   "Carrier_67_SitopSelectStatus" AT %I3716.3 : Bool;   // SITOP SELECT STATUS
   "Carrier_67_DCsupplyOnPSCB2" AT %I3716.4 : Bool;   // DC SUPPLY ON PSCB 2
   "Carrier_67_SpareInput(4_5)" AT %I3716.5 : Bool;   // SPARE INPUT
   "Carrier_67_SpareInput(4_6)" AT %I3716.6 : Bool;   // SPARE INPUT
   "Carrier_67_SpareInput(4_7)" AT %I3716.7 : Bool;   // SPARE INPUT
   "Carrier_67_PB1_ProdHoldLH" AT %I3717.0 : Bool;   // PB 1 PRODUCTION HOLD LH
   "Carrier_67_PB2_ResetLH" AT %I3717.1 : Bool;   // PB 2 RESET LH
   "Carrier_67_PB3_ProdHoldRH" AT %I3717.2 : Bool;   // PB 3 PRODUCTION HOLD RH
   "Carrier_67_PB4_ResetRH" AT %I3717.3 : Bool;   // PB 4 RESET RH
   "Carrier_67_SpareInput(4_14)" AT %I3717.4 : Bool;   // SPARE INPUT
   "Carrier_67_SpareInput(4_15)" AT %I3717.5 : Bool;   // SPARE INPUT
   "Carrier_67_SpareInput(4_16)" AT %I3717.6 : Bool;   // SPARE INPUT
   "Carrier_67_SpareInput(4_17)" AT %I3717.7 : Bool;   // SPARE INPUT
   "Carrier_67_Slot5_Output" AT %IW3718 : Word;   // SLOT 5 OUTPUT WORD
   "Carrier_67_IRD400_HMI_24VDC_ENABLE" AT %I3718.0 : Bool;   // IRD 400 PANEL HMI 24V DC POWER
   "Carrier_67_FaultLight_LH" AT %I3718.1 : Bool;   // FAULT LIGHT LH
   "Carrier_67_RunLight_LH" AT %I3718.2 : Bool;   // RUN LIGHT LH
   "Carrier_67_FaultLight_RH" AT %I3718.3 : Bool;   // FAULT LIGHT RH
   "Carrier_67_RunLight_RH" AT %I3718.4 : Bool;   // RUN LIGHT RH
   "Carrier_67_SpareOutput(5_5)" AT %I3718.5 : Bool;   // SPARE OUTPUT
   "Carrier_67_SpareOutput(5_6)" AT %I3718.6 : Bool;   // SPARE OUTPUT
   "Carrier_67_SpareOutput(5_7)" AT %I3718.7 : Bool;   // SPARE OUTPUT
   "Carrier_67_ActualSpeed" AT %IW3720 : Word;   // ACTUAL SPEED
   "Carrier_67_CarrierDriveAlarm" AT %IW3722 : Word;   // CARRIER DRIVE ALARM
   "Carrier_67_CarrierDriveWarning" AT %IW3724 : Word;   // CARRIER DRIVE WARNING
   "Carrier_68_Status" AT %IW3750 : Word;   // CARRIER STATUS WORD
   "Carrier_68_Status.0" AT %I3750.0 : Bool;   // HEARTBEAT
   "Carrier_68_Status.1" AT %I3750.1 : Bool;   // MANUAL
   "Carrier_68_Status.2" AT %I3750.2 : Bool;   // IN_AUTO
   "Carrier_68_Status.3" AT %I3750.3 : Bool;   // POSITIONING_COMPLETE
   "Carrier_68_Status.4" AT %I3750.4 : Bool;   // PRODUCTION HOLD
   "Carrier_68_Status.5" AT %I3750.5 : Bool;   // CARRIER MOVING FORWARD
   "Carrier_68_Status.6" AT %I3750.6 : Bool;   // CARRIER MOVING REVERSE
   "Carrier_68_Status.7" AT %I3750.7 : Bool;   // CARRIER FAULT
   "Carrier_68_Status.8" AT %I3751.0 : Bool;   // CRASH DETECT TRIPPED
   "Carrier_68_Status.9" AT %I3751.1 : Bool;
   "Carrier_68_Status.10" AT %I3751.2 : Bool;
   "Carrier_68_Status.11" AT %I3751.3 : Bool;
   "Carrier_68_Status.12" AT %I3751.4 : Bool;
   "Carrier_68_Status.13" AT %I3751.5 : Bool;
   "Carrier_68_Status.14" AT %I3751.6 : Bool;
   "Carrier_68_Status.15" AT %I3751.7 : Bool;
   "Carrier_68_SDCFaultCode" AT %IW3752 : Word;   // SDC FAULT CODE
   "Carrier_68_CarrierPosition" AT %ID3754 : DWord;   // CARRIER POSITION
   "Carrier_68_CarrierNumber" AT %IW3758 : Word;   // CARRIER NUMBER
   "Carrier_68_G120DControlWord" AT %IW3760 : Word;   // G120D_STW1_CONTROL
   "Carrier_68_G120DControlWord.0" AT %I3760.0 : Bool;   // Bit_00_ON
   "Carrier_68_G120DControlWord.1" AT %I3760.1 : Bool;   // Bit_01_AUS2_INH
   "Carrier_68_G120DControlWord.2" AT %I3760.2 : Bool;   // Bit_02_AUS3_STOP
   "Carrier_68_G120DControlWord.3" AT %I3760.3 : Bool;   // Bit_03_EN
   "Carrier_68_G120DControlWord.4" AT %I3760.4 : Bool;   // Bit_04_EN_RAMP
   "Carrier_68_G120DControlWord.5" AT %I3760.5 : Bool;   // Bit_05_START_RAMP
   "Carrier_68_G120DControlWord.6" AT %I3760.6 : Bool;   // Bit_06_SETPOINT
   "Carrier_68_G120DControlWord.7" AT %I3760.7 : Bool;   // Bit_07_RESET
   "Carrier_68_G120DControlWord.8" AT %I3761.0 : Bool;   // Bit_08_JOG_R
   "Carrier_68_G120DControlWord.9" AT %I3761.1 : Bool;   // Bit_09_JOG_L
   "Carrier_68_G120DControlWord.10" AT %I3761.2 : Bool;   // Bit_10_CONTR_PLC
   "Carrier_68_G120DControlWord.11" AT %I3761.3 : Bool;   // Bit_11_REVERSE
   "Carrier_68_G120DControlWord.12" AT %I3761.4 : Bool;   // Bit_12_BRAKE_RELEASE
   "Carrier_68_G120DControlWord.13" AT %I3761.5 : Bool;   // Bit_13_DDS
   "Carrier_68_G120DControlWord.14" AT %I3761.6 : Bool;   // Bit_14_DO0
   "Carrier_68_G120DControlWord.15" AT %I3761.7 : Bool;   // Bit_15_DO1
   "Carrier_68_G120DStatusWord" AT %IW3762 : Word;   // G120D_ZSW1_STATUS
   "Carrier_68_G120DStatusWord.0" AT %I3762.0 : Bool;   // Bit_00_READY_RUN
   "Carrier_68_G120DStatusWord.1" AT %I3762.1 : Bool;   // Bit_01_READY_ON
   "Carrier_68_G120DStatusWord.2" AT %I3762.2 : Bool;   // Bit_02_ENABLE
   "Carrier_68_G120DStatusWord.3" AT %I3762.3 : Bool;   // Bit_03_FAULT
   "Carrier_68_G120DStatusWord.4" AT %I3762.4 : Bool;   // Bit_04_OFF2
   "Carrier_68_G120DStatusWord.5" AT %I3762.5 : Bool;   // Bit_05_OFF3
   "Carrier_68_G120DStatusWord.6" AT %I3762.6 : Bool;   // Bit_06_LOCK_OUT
   "Carrier_68_G120DStatusWord.7" AT %I3762.7 : Bool;   // Bit_07_WARN
   "Carrier_68_G120DStatusWord.8" AT %I3763.0 : Bool;   // Bit_08_NO_DEVIATION
   "Carrier_68_G120DStatusWord.9" AT %I3763.1 : Bool;   // Bit_09_CONTR_PLC
   "Carrier_68_G120DStatusWord.10" AT %I3763.2 : Bool;   // Bit_10_F_MAX
   "Carrier_68_G120DStatusWord.11" AT %I3763.3 : Bool;   // Bit_11_LIMIT_REACHED
   "Carrier_68_G120DStatusWord.12" AT %I3763.4 : Bool;   // Bit_12_BRAKE_OPEN
   "Carrier_68_G120DStatusWord.13" AT %I3763.5 : Bool;   // Bit_13_NO_OVERTEMP
   "Carrier_68_G120DStatusWord.14" AT %I3763.6 : Bool;   // Bit_14_CW_CCW
   "Carrier_68_G120DStatusWord.15" AT %I3763.7 : Bool;   // Bit_15_OVERL
   "Carrier_68_Slot2_Input" AT %IW3764 : Word;   // SLOT 2 INPUT WORD
   "Carrier_68_CrashDetectSW" AT %I3764.0 : Bool;   // CRASH DETECT SW
   "Carrier_68_SpareSafetyInput(2_1)" AT %I3764.1 : Bool;   // SPARE SAFETY INPUT
   "Carrier_68_SpareSafetyInput(2_2)" AT %I3764.2 : Bool;   // SPARE SAFETY INPUT
   "Carrier_68_SpareSafetyInput(2_3)" AT %I3764.3 : Bool;   // SPARE SAFETY INPUT
   "Carrier_68_SpareSafetyInput(2_4)" AT %I3764.4 : Bool;   // SPARE SAFETY INPUT
   "Carrier_68_SpareSafetyInput(2_5)" AT %I3764.5 : Bool;   // SPARE SAFETY INPUT
   "Carrier_68_SpareSafetyInput(2_6)" AT %I3764.6 : Bool;   // SPARE SAFETY INPUT
   "Carrier_68_SpareSafetyInput(2_7)" AT %I3764.7 : Bool;   // SPARE SAFETY INPUT
   "Carrier_68_Slot3_SafetyOutput" AT %IW3765 : Word;   // SLOT 3 SAFETY OUTPUT WORD
   "Carrier_68_Crash_Detect_OK" AT %I3765.0 : Bool;   // CARRIER CRASH DETECT
   "Carrier_68_SpareSafetyOutput(3_1)" AT %I3765.1 : Bool;   // SPARE SAFETY OUTPUT
   "Carrier_68_SpareSafetyOutput(3_2)" AT %I3765.2 : Bool;   // SPARE SAFETY OUTPUT
   "Carrier_68_SpareSafetyOutput(3_3)" AT %I3765.3 : Bool;   // SPARE SAFETY OUTPUT
   "Carrier_68_SpareSafetyOutput(3_4)" AT %I3765.4 : Bool;   // SPARE SAFETY OUTPUT
   "Carrier_68_SpareSafetyOutput(3_5)" AT %I3765.5 : Bool;   // SPARE SAFETY OUTPUT
   "Carrier_68_SpareSafetyOutput(3_6)" AT %I3765.6 : Bool;   // SPARE SAFETY OUTPUT
   "Carrier_68_SpareSafetyOutput(3_7)" AT %I3765.7 : Bool;   // SPARE SAFETY OUTPUT
   "Carrier_68_Slot4_Input" AT %IW3766 : Word;   // SLOT 4 INPUT WORD
   "Carrier_68_480VPowerOn_MDCB1" AT %I3766.0 : Bool;   // 480 VAC POWER ON MDCB 1
   "Carrier_68_SpareInput(4_1)" AT %I3766.1 : Bool;   // SPARE INPUT
   "Carrier_68_SpareInput(4_2)" AT %I3766.2 : Bool;   // SPARE INPUT
   "Carrier_68_SitopSelectStatus" AT %I3766.3 : Bool;   // SITOP SELECT STATUS
   "Carrier_68_DCsupplyOnPSCB2" AT %I3766.4 : Bool;   // DC SUPPLY ON PSCB 2
   "Carrier_68_SpareInput(4_5)" AT %I3766.5 : Bool;   // SPARE INPUT
   "Carrier_68_SpareInput(4_6)" AT %I3766.6 : Bool;   // SPARE INPUT
   "Carrier_68_SpareInput(4_7)" AT %I3766.7 : Bool;   // SPARE INPUT
   "Carrier_68_PB1_ProdHoldLH" AT %I3767.0 : Bool;   // PB 1 PRODUCTION HOLD LH
   "Carrier_68_PB2_ResetLH" AT %I3767.1 : Bool;   // PB 2 RESET LH
   "Carrier_68_PB3_ProdHoldRH" AT %I3767.2 : Bool;   // PB 3 PRODUCTION HOLD RH
   "Carrier_68_PB4_ResetRH" AT %I3767.3 : Bool;   // PB 4 RESET RH
   "Carrier_68_SpareInput(4_14)" AT %I3767.4 : Bool;   // SPARE INPUT
   "Carrier_68_SpareInput(4_15)" AT %I3767.5 : Bool;   // SPARE INPUT
   "Carrier_68_SpareInput(4_16)" AT %I3767.6 : Bool;   // SPARE INPUT
   "Carrier_68_SpareInput(4_17)" AT %I3767.7 : Bool;   // SPARE INPUT
   "Carrier_68_Slot5_Output" AT %IW3768 : Word;   // SLOT 5 OUTPUT WORD
   "Carrier_68_IRD400_HMI_24VDC_ENABLE" AT %I3768.0 : Bool;   // IRD 400 PANEL HMI 24V DC POWER
   "Carrier_68_FaultLight_LH" AT %I3768.1 : Bool;   // FAULT LIGHT LH
   "Carrier_68_RunLight_LH" AT %I3768.2 : Bool;   // RUN LIGHT LH
   "Carrier_68_FaultLight_RH" AT %I3768.3 : Bool;   // FAULT LIGHT RH
   "Carrier_68_RunLight_RH" AT %I3768.4 : Bool;   // RUN LIGHT RH
   "Carrier_68_SpareOutput(5_5)" AT %I3768.5 : Bool;   // SPARE OUTPUT
   "Carrier_68_SpareOutput(5_6)" AT %I3768.6 : Bool;   // SPARE OUTPUT
   "Carrier_68_SpareOutput(5_7)" AT %I3768.7 : Bool;   // SPARE OUTPUT
   "Carrier_68_ActualSpeed" AT %IW3770 : Word;   // ACTUAL SPEED
   "Carrier_68_CarrierDriveAlarm" AT %IW3772 : Word;   // CARRIER DRIVE ALARM
   "Carrier_68_CarrierDriveWarning" AT %IW3774 : Word;   // CARRIER DRIVE WARNING
   "Carrier_69_Status" AT %IW3800 : Word;   // CARRIER STATUS WORD
   "Carrier_69_Status.0" AT %I3800.0 : Bool;   // HEARTBEAT
   "Carrier_69_Status.1" AT %I3800.1 : Bool;   // MANUAL
   "Carrier_69_Status.2" AT %I3800.2 : Bool;   // IN_AUTO
   "Carrier_69_Status.3" AT %I3800.3 : Bool;   // POSITIONING_COMPLETE
   "Carrier_69_Status.4" AT %I3800.4 : Bool;   // PRODUCTION HOLD
   "Carrier_69_Status.5" AT %I3800.5 : Bool;   // CARRIER MOVING FORWARD
   "Carrier_69_Status.6" AT %I3800.6 : Bool;   // CARRIER MOVING REVERSE
   "Carrier_69_Status.7" AT %I3800.7 : Bool;   // CARRIER FAULT
   "Carrier_69_Status.8" AT %I3801.0 : Bool;   // CRASH DETECT TRIPPED
   "Carrier_69_Status.9" AT %I3801.1 : Bool;
   "Carrier_69_Status.10" AT %I3801.2 : Bool;
   "Carrier_69_Status.11" AT %I3801.3 : Bool;
   "Carrier_69_Status.12" AT %I3801.4 : Bool;
   "Carrier_69_Status.13" AT %I3801.5 : Bool;
   "Carrier_69_Status.14" AT %I3801.6 : Bool;
   "Carrier_69_Status.15" AT %I3801.7 : Bool;
   "Carrier_69_SDCFaultCode" AT %IW3802 : Word;   // SDC FAULT CODE
   "Carrier_69_CarrierPosition" AT %ID3804 : DWord;   // CARRIER POSITION
   "Carrier_69_CarrierNumber" AT %IW3808 : Word;   // CARRIER NUMBER
   "Carrier_69_G120DControlWord" AT %IW3810 : Word;   // G120D_STW1_CONTROL
   "Carrier_69_G120DControlWord.0" AT %I3810.0 : Bool;   // Bit_00_ON
   "Carrier_69_G120DControlWord.1" AT %I3810.1 : Bool;   // Bit_01_AUS2_INH
   "Carrier_69_G120DControlWord.2" AT %I3810.2 : Bool;   // Bit_02_AUS3_STOP
   "Carrier_69_G120DControlWord.3" AT %I3810.3 : Bool;   // Bit_03_EN
   "Carrier_69_G120DControlWord.4" AT %I3810.4 : Bool;   // Bit_04_EN_RAMP
   "Carrier_69_G120DControlWord.5" AT %I3810.5 : Bool;   // Bit_05_START_RAMP
   "Carrier_69_G120DControlWord.6" AT %I3810.6 : Bool;   // Bit_06_SETPOINT
   "Carrier_69_G120DControlWord.7" AT %I3810.7 : Bool;   // Bit_07_RESET
   "Carrier_69_G120DControlWord.8" AT %I3811.0 : Bool;   // Bit_08_JOG_R
   "Carrier_69_G120DControlWord.9" AT %I3811.1 : Bool;   // Bit_09_JOG_L
   "Carrier_69_G120DControlWord.10" AT %I3811.2 : Bool;   // Bit_10_CONTR_PLC
   "Carrier_69_G120DControlWord.11" AT %I3811.3 : Bool;   // Bit_11_REVERSE
   "Carrier_69_G120DControlWord.12" AT %I3811.4 : Bool;   // Bit_12_BRAKE_RELEASE
   "Carrier_69_G120DControlWord.13" AT %I3811.5 : Bool;   // Bit_13_DDS
   "Carrier_69_G120DControlWord.14" AT %I3811.6 : Bool;   // Bit_14_DO0
   "Carrier_69_G120DControlWord.15" AT %I3811.7 : Bool;   // Bit_15_DO1
   "Carrier_69_G120DStatusWord" AT %IW3812 : Word;   // G120D_ZSW1_STATUS
   "Carrier_69_G120DStatusWord.0" AT %I3812.0 : Bool;   // Bit_00_READY_RUN
   "Carrier_69_G120DStatusWord.1" AT %I3812.1 : Bool;   // Bit_01_READY_ON
   "Carrier_69_G120DStatusWord.2" AT %I3812.2 : Bool;   // Bit_02_ENABLE
   "Carrier_69_G120DStatusWord.3" AT %I3812.3 : Bool;   // Bit_03_FAULT
   "Carrier_69_G120DStatusWord.4" AT %I3812.4 : Bool;   // Bit_04_OFF2
   "Carrier_69_G120DStatusWord.5" AT %I3812.5 : Bool;   // Bit_05_OFF3
   "Carrier_69_G120DStatusWord.6" AT %I3812.6 : Bool;   // Bit_06_LOCK_OUT
   "Carrier_69_G120DStatusWord.7" AT %I3812.7 : Bool;   // Bit_07_WARN
   "Carrier_69_G120DStatusWord.8" AT %I3813.0 : Bool;   // Bit_08_NO_DEVIATION
   "Carrier_69_G120DStatusWord.9" AT %I3813.1 : Bool;   // Bit_09_CONTR_PLC
   "Carrier_69_G120DStatusWord.10" AT %I3813.2 : Bool;   // Bit_10_F_MAX
   "Carrier_69_G120DStatusWord.11" AT %I3813.3 : Bool;   // Bit_11_LIMIT_REACHED
   "Carrier_69_G120DStatusWord.12" AT %I3813.4 : Bool;   // Bit_12_BRAKE_OPEN
   "Carrier_69_G120DStatusWord.13" AT %I3813.5 : Bool;   // Bit_13_NO_OVERTEMP
   "Carrier_69_G120DStatusWord.14" AT %I3813.6 : Bool;   // Bit_14_CW_CCW
   "Carrier_69_G120DStatusWord.15" AT %I3813.7 : Bool;   // Bit_15_OVERL
   "Carrier_69_Slot2_Input" AT %IW3814 : Word;   // SLOT 2 INPUT WORD
   "Carrier_69_CrashDetectSW" AT %I3814.0 : Bool;   // CRASH DETECT SW
   "Carrier_69_SpareSafetyInput(2_1)" AT %I3814.1 : Bool;   // SPARE SAFETY INPUT
   "Carrier_69_SpareSafetyInput(2_2)" AT %I3814.2 : Bool;   // SPARE SAFETY INPUT
   "Carrier_69_SpareSafetyInput(2_3)" AT %I3814.3 : Bool;   // SPARE SAFETY INPUT
   "Carrier_69_SpareSafetyInput(2_4)" AT %I3814.4 : Bool;   // SPARE SAFETY INPUT
   "Carrier_69_SpareSafetyInput(2_5)" AT %I3814.5 : Bool;   // SPARE SAFETY INPUT
   "Carrier_69_SpareSafetyInput(2_6)" AT %I3814.6 : Bool;   // SPARE SAFETY INPUT
   "Carrier_69_SpareSafetyInput(2_7)" AT %I3814.7 : Bool;   // SPARE SAFETY INPUT
   "Carrier_69_Slot3_SafetyOutput" AT %IW3815 : Word;   // SLOT 3 SAFETY OUTPUT WORD
   "Carrier_69_Crash_Detect_OK" AT %I3815.0 : Bool;   // CARRIER CRASH DETECT
   "Carrier_69_SpareSafetyOutput(3_1)" AT %I3815.1 : Bool;   // SPARE SAFETY OUTPUT
   "Carrier_69_SpareSafetyOutput(3_2)" AT %I3815.2 : Bool;   // SPARE SAFETY OUTPUT
   "Carrier_69_SpareSafetyOutput(3_3)" AT %I3815.3 : Bool;   // SPARE SAFETY OUTPUT
   "Carrier_69_SpareSafetyOutput(3_4)" AT %I3815.4 : Bool;   // SPARE SAFETY OUTPUT
   "Carrier_69_SpareSafetyOutput(3_5)" AT %I3815.5 : Bool;   // SPARE SAFETY OUTPUT
   "Carrier_69_SpareSafetyOutput(3_6)" AT %I3815.6 : Bool;   // SPARE SAFETY OUTPUT
   "Carrier_69_SpareSafetyOutput(3_7)" AT %I3815.7 : Bool;   // SPARE SAFETY OUTPUT
   "Carrier_69_Slot4_Input" AT %IW3816 : Word;   // SLOT 4 INPUT WORD
   "Carrier_69_480VPowerOn_MDCB1" AT %I3816.0 : Bool;   // 480 VAC POWER ON MDCB 1
   "Carrier_69_SpareInput(4_1)" AT %I3816.1 : Bool;   // SPARE INPUT
   "Carrier_69_SpareInput(4_2)" AT %I3816.2 : Bool;   // SPARE INPUT
   "Carrier_69_SitopSelectStatus" AT %I3816.3 : Bool;   // SITOP SELECT STATUS
   "Carrier_69_DCsupplyOnPSCB2" AT %I3816.4 : Bool;   // DC SUPPLY ON PSCB 2
   "Carrier_69_SpareInput(4_5)" AT %I3816.5 : Bool;   // SPARE INPUT
   "Carrier_69_SpareInput(4_6)" AT %I3816.6 : Bool;   // SPARE INPUT
   "Carrier_69_SpareInput(4_7)" AT %I3816.7 : Bool;   // SPARE INPUT
   "Carrier_69_PB1_ProdHoldLH" AT %I3817.0 : Bool;   // PB 1 PRODUCTION HOLD LH
   "Carrier_69_PB2_ResetLH" AT %I3817.1 : Bool;   // PB 2 RESET LH
   "Carrier_69_PB3_ProdHoldRH" AT %I3817.2 : Bool;   // PB 3 PRODUCTION HOLD RH
   "Carrier_69_PB4_ResetRH" AT %I3817.3 : Bool;   // PB 4 RESET RH
   "Carrier_69_SpareInput(4_14)" AT %I3817.4 : Bool;   // SPARE INPUT
   "Carrier_69_SpareInput(4_15)" AT %I3817.5 : Bool;   // SPARE INPUT
   "Carrier_69_SpareInput(4_16)" AT %I3817.6 : Bool;   // SPARE INPUT
   "Carrier_69_SpareInput(4_17)" AT %I3817.7 : Bool;   // SPARE INPUT
   "Carrier_69_Slot5_Output" AT %IW3818 : Word;   // SLOT 5 OUTPUT WORD
   "Carrier_69_IRD400_HMI_24VDC_ENABLE" AT %I3818.0 : Bool;   // IRD 400 PANEL HMI 24V DC POWER
   "Carrier_69_FaultLight_LH" AT %I3818.1 : Bool;   // FAULT LIGHT LH
   "Carrier_69_RunLight_LH" AT %I3818.2 : Bool;   // RUN LIGHT LH
   "Carrier_69_FaultLight_RH" AT %I3818.3 : Bool;   // FAULT LIGHT RH
   "Carrier_69_RunLight_RH" AT %I3818.4 : Bool;   // RUN LIGHT RH
   "Carrier_69_SpareOutput(5_5)" AT %I3818.5 : Bool;   // SPARE OUTPUT
   "Carrier_69_SpareOutput(5_6)" AT %I3818.6 : Bool;   // SPARE OUTPUT
   "Carrier_69_SpareOutput(5_7)" AT %I3818.7 : Bool;   // SPARE OUTPUT
   "Carrier_69_ActualSpeed" AT %IW3820 : Word;   // ACTUAL SPEED
   "Carrier_69_CarrierDriveAlarm" AT %IW3822 : Word;   // CARRIER DRIVE ALARM
   "Carrier_69_CarrierDriveWarning" AT %IW3824 : Word;   // CARRIER DRIVE WARNING
   "Carrier_70_Status" AT %IW3850 : Word;   // CARRIER STATUS WORD
   "Carrier_70_Status.0" AT %I3850.0 : Bool;   // HEARTBEAT
   "Carrier_70_Status.1" AT %I3850.1 : Bool;   // MANUAL
   "Carrier_70_Status.2" AT %I3850.2 : Bool;   // IN_AUTO
   "Carrier_70_Status.3" AT %I3850.3 : Bool;   // POSITIONING_COMPLETE
   "Carrier_70_Status.4" AT %I3850.4 : Bool;   // PRODUCTION HOLD
   "Carrier_70_Status.5" AT %I3850.5 : Bool;   // CARRIER MOVING FORWARD
   "Carrier_70_Status.6" AT %I3850.6 : Bool;   // CARRIER MOVING REVERSE
   "Carrier_70_Status.7" AT %I3850.7 : Bool;   // CARRIER FAULT
   "Carrier_70_Status.8" AT %I3851.0 : Bool;   // CRASH DETECT TRIPPED
   "Carrier_70_Status.9" AT %I3851.1 : Bool;
   "Carrier_70_Status.10" AT %I3851.2 : Bool;
   "Carrier_70_Status.11" AT %I3851.3 : Bool;
   "Carrier_70_Status.12" AT %I3851.4 : Bool;
   "Carrier_70_Status.13" AT %I3851.5 : Bool;
   "Carrier_70_Status.14" AT %I3851.6 : Bool;
   "Carrier_70_Status.15" AT %I3851.7 : Bool;
   "Carrier_70_SDCFaultCode" AT %IW3852 : Word;   // SDC FAULT CODE
   "Carrier_70_CarrierPosition" AT %ID3854 : DWord;   // CARRIER POSITION
   "Carrier_70_CarrierNumber" AT %IW3858 : Word;   // CARRIER NUMBER
   "Carrier_70_G120DControlWord" AT %IW3860 : Word;   // G120D_STW1_CONTROL
   "Carrier_70_G120DControlWord.0" AT %I3860.0 : Bool;   // Bit_00_ON
   "Carrier_70_G120DControlWord.1" AT %I3860.1 : Bool;   // Bit_01_AUS2_INH
   "Carrier_70_G120DControlWord.2" AT %I3860.2 : Bool;   // Bit_02_AUS3_STOP
   "Carrier_70_G120DControlWord.3" AT %I3860.3 : Bool;   // Bit_03_EN
   "Carrier_70_G120DControlWord.4" AT %I3860.4 : Bool;   // Bit_04_EN_RAMP
   "Carrier_70_G120DControlWord.5" AT %I3860.5 : Bool;   // Bit_05_START_RAMP
   "Carrier_70_G120DControlWord.6" AT %I3860.6 : Bool;   // Bit_06_SETPOINT
   "Carrier_70_G120DControlWord.7" AT %I3860.7 : Bool;   // Bit_07_RESET
   "Carrier_70_G120DControlWord.8" AT %I3861.0 : Bool;   // Bit_08_JOG_R
   "Carrier_70_G120DControlWord.9" AT %I3861.1 : Bool;   // Bit_09_JOG_L
   "Carrier_70_G120DControlWord.10" AT %I3861.2 : Bool;   // Bit_10_CONTR_PLC
   "Carrier_70_G120DControlWord.11" AT %I3861.3 : Bool;   // Bit_11_REVERSE
   "Carrier_70_G120DControlWord.12" AT %I3861.4 : Bool;   // Bit_12_BRAKE_RELEASE
   "Carrier_70_G120DControlWord.13" AT %I3861.5 : Bool;   // Bit_13_DDS
   "Carrier_70_G120DControlWord.14" AT %I3861.6 : Bool;   // Bit_14_DO0
   "Carrier_70_G120DControlWord.15" AT %I3861.7 : Bool;   // Bit_15_DO1
   "Carrier_70_G120DStatusWord" AT %IW3862 : Word;   // G120D_ZSW1_STATUS
   "Carrier_70_G120DStatusWord.0" AT %I3862.0 : Bool;   // Bit_00_READY_RUN
   "Carrier_70_G120DStatusWord.1" AT %I3862.1 : Bool;   // Bit_01_READY_ON
   "Carrier_70_G120DStatusWord.2" AT %I3862.2 : Bool;   // Bit_02_ENABLE
   "Carrier_70_G120DStatusWord.3" AT %I3862.3 : Bool;   // Bit_03_FAULT
   "Carrier_70_G120DStatusWord.4" AT %I3862.4 : Bool;   // Bit_04_OFF2
   "Carrier_70_G120DStatusWord.5" AT %I3862.5 : Bool;   // Bit_05_OFF3
   "Carrier_70_G120DStatusWord.6" AT %I3862.6 : Bool;   // Bit_06_LOCK_OUT
   "Carrier_70_G120DStatusWord.7" AT %I3862.7 : Bool;   // Bit_07_WARN
   "Carrier_70_G120DStatusWord.8" AT %I3863.0 : Bool;   // Bit_08_NO_DEVIATION
   "Carrier_70_G120DStatusWord.9" AT %I3863.1 : Bool;   // Bit_09_CONTR_PLC
   "Carrier_70_G120DStatusWord.10" AT %I3863.2 : Bool;   // Bit_10_F_MAX
   "Carrier_70_G120DStatusWord.11" AT %I3863.3 : Bool;   // Bit_11_LIMIT_REACHED
   "Carrier_70_G120DStatusWord.12" AT %I3863.4 : Bool;   // Bit_12_BRAKE_OPEN
   "Carrier_70_G120DStatusWord.13" AT %I3863.5 : Bool;   // Bit_13_NO_OVERTEMP
   "Carrier_70_G120DStatusWord.14" AT %I3863.6 : Bool;   // Bit_14_CW_CCW
   "Carrier_70_G120DStatusWord.15" AT %I3863.7 : Bool;   // Bit_15_OVERL
   "Carrier_70_Slot2_Input" AT %IW3864 : Word;   // SLOT 2 INPUT WORD
   "Carrier_70_CrashDetectSW" AT %I3864.0 : Bool;   // CRASH DETECT SW
   "Carrier_70_SpareSafetyInput(2_1)" AT %I3864.1 : Bool;   // SPARE SAFETY INPUT
   "Carrier_70_SpareSafetyInput(2_2)" AT %I3864.2 : Bool;   // SPARE SAFETY INPUT
   "Carrier_70_SpareSafetyInput(2_3)" AT %I3864.3 : Bool;   // SPARE SAFETY INPUT
   "Carrier_70_SpareSafetyInput(2_4)" AT %I3864.4 : Bool;   // SPARE SAFETY INPUT
   "Carrier_70_SpareSafetyInput(2_5)" AT %I3864.5 : Bool;   // SPARE SAFETY INPUT
   "Carrier_70_SpareSafetyInput(2_6)" AT %I3864.6 : Bool;   // SPARE SAFETY INPUT
   "Carrier_70_SpareSafetyInput(2_7)" AT %I3864.7 : Bool;   // SPARE SAFETY INPUT
   "Carrier_70_Slot3_SafetyOutput" AT %IW3865 : Word;   // SLOT 3 SAFETY OUTPUT WORD
   "Carrier_70_Crash_Detect_OK" AT %I3865.0 : Bool;   // CARRIER CRASH DETECT
   "Carrier_70_SpareSafetyOutput(3_1)" AT %I3865.1 : Bool;   // SPARE SAFETY OUTPUT
   "Carrier_70_SpareSafetyOutput(3_2)" AT %I3865.2 : Bool;   // SPARE SAFETY OUTPUT
   "Carrier_70_SpareSafetyOutput(3_3)" AT %I3865.3 : Bool;   // SPARE SAFETY OUTPUT
   "Carrier_70_SpareSafetyOutput(3_4)" AT %I3865.4 : Bool;   // SPARE SAFETY OUTPUT
   "Carrier_70_SpareSafetyOutput(3_5)" AT %I3865.5 : Bool;   // SPARE SAFETY OUTPUT
   "Carrier_70_SpareSafetyOutput(3_6)" AT %I3865.6 : Bool;   // SPARE SAFETY OUTPUT
   "Carrier_70_SpareSafetyOutput(3_7)" AT %I3865.7 : Bool;   // SPARE SAFETY OUTPUT
   "Carrier_70_Slot4_Input" AT %IW3866 : Word;   // SLOT 4 INPUT WORD
   "Carrier_70_480VPowerOn_MDCB1" AT %I3866.0 : Bool;   // 480 VAC POWER ON MDCB 1
   "Carrier_70_SpareInput(4_1)" AT %I3866.1 : Bool;   // SPARE INPUT
   "Carrier_70_SpareInput(4_2)" AT %I3866.2 : Bool;   // SPARE INPUT
   "Carrier_70_SitopSelectStatus" AT %I3866.3 : Bool;   // SITOP SELECT STATUS
   "Carrier_70_DCsupplyOnPSCB2" AT %I3866.4 : Bool;   // DC SUPPLY ON PSCB 2
   "Carrier_70_SpareInput(4_5)" AT %I3866.5 : Bool;   // SPARE INPUT
   "Carrier_70_SpareInput(4_6)" AT %I3866.6 : Bool;   // SPARE INPUT
   "Carrier_70_SpareInput(4_7)" AT %I3866.7 : Bool;   // SPARE INPUT
   "Carrier_70_PB1_ProdHoldLH" AT %I3867.0 : Bool;   // PB 1 PRODUCTION HOLD LH
   "Carrier_70_PB2_ResetLH" AT %I3867.1 : Bool;   // PB 2 RESET LH
   "Carrier_70_PB3_ProdHoldRH" AT %I3867.2 : Bool;   // PB 3 PRODUCTION HOLD RH
   "Carrier_70_PB4_ResetRH" AT %I3867.3 : Bool;   // PB 4 RESET RH
   "Carrier_70_SpareInput(4_14)" AT %I3867.4 : Bool;   // SPARE INPUT
   "Carrier_70_SpareInput(4_15)" AT %I3867.5 : Bool;   // SPARE INPUT
   "Carrier_70_SpareInput(4_16)" AT %I3867.6 : Bool;   // SPARE INPUT
   "Carrier_70_SpareInput(4_17)" AT %I3867.7 : Bool;   // SPARE INPUT
   "Carrier_70_Slot5_Output" AT %IW3868 : Word;   // SLOT 5 OUTPUT WORD
   "Carrier_70_IRD400_HMI_24VDC_ENABLE" AT %I3868.0 : Bool;   // IRD 400 PANEL HMI 24V DC POWER
   "Carrier_70_FaultLight_LH" AT %I3868.1 : Bool;   // FAULT LIGHT LH
   "Carrier_70_RunLight_LH" AT %I3868.2 : Bool;   // RUN LIGHT LH
   "Carrier_70_FaultLight_RH" AT %I3868.3 : Bool;   // FAULT LIGHT RH
   "Carrier_70_RunLight_RH" AT %I3868.4 : Bool;   // RUN LIGHT RH
   "Carrier_70_SpareOutput(5_5)" AT %I3868.5 : Bool;   // SPARE OUTPUT
   "Carrier_70_SpareOutput(5_6)" AT %I3868.6 : Bool;   // SPARE OUTPUT
   "Carrier_70_SpareOutput(5_7)" AT %I3868.7 : Bool;   // SPARE OUTPUT
   "Carrier_70_ActualSpeed" AT %IW3870 : Word;   // ACTUAL SPEED
   "Carrier_70_CarrierDriveAlarm" AT %IW3872 : Word;   // CARRIER DRIVE ALARM
   "Carrier_70_CarrierDriveWarning" AT %IW3874 : Word;   // CARRIER DRIVE WARNING
   "Carrier_71_Status" AT %IW3900 : Word;   // CARRIER STATUS WORD
   "Carrier_71_Status.0" AT %I3900.0 : Bool;   // HEARTBEAT
   "Carrier_71_Status.1" AT %I3900.1 : Bool;   // MANUAL
   "Carrier_71_Status.2" AT %I3900.2 : Bool;   // IN_AUTO
   "Carrier_71_Status.3" AT %I3900.3 : Bool;   // POSITIONING_COMPLETE
   "Carrier_71_Status.4" AT %I3900.4 : Bool;   // PRODUCTION HOLD
   "Carrier_71_Status.5" AT %I3900.5 : Bool;   // CARRIER MOVING FORWARD
   "Carrier_71_Status.6" AT %I3900.6 : Bool;   // CARRIER MOVING REVERSE
   "Carrier_71_Status.7" AT %I3900.7 : Bool;   // CARRIER FAULT
   "Carrier_71_Status.8" AT %I3901.0 : Bool;   // CRASH DETECT TRIPPED
   "Carrier_71_Status.9" AT %I3901.1 : Bool;
   "Carrier_71_Status.10" AT %I3901.2 : Bool;
   "Carrier_71_Status.11" AT %I3901.3 : Bool;
   "Carrier_71_Status.12" AT %I3901.4 : Bool;
   "Carrier_71_Status.13" AT %I3901.5 : Bool;
   "Carrier_71_Status.14" AT %I3901.6 : Bool;
   "Carrier_71_Status.15" AT %I3901.7 : Bool;
   "Carrier_71_SDCFaultCode" AT %IW3902 : Word;   // SDC FAULT CODE
   "Carrier_71_CarrierPosition" AT %ID3904 : DWord;   // CARRIER POSITION
   "Carrier_71_CarrierNumber" AT %IW3908 : Word;   // CARRIER NUMBER
   "Carrier_71_G120DControlWord" AT %IW3910 : Word;   // G120D_STW1_CONTROL
   "Carrier_71_G120DControlWord.0" AT %I3910.0 : Bool;   // Bit_00_ON
   "Carrier_71_G120DControlWord.1" AT %I3910.1 : Bool;   // Bit_01_AUS2_INH
   "Carrier_71_G120DControlWord.2" AT %I3910.2 : Bool;   // Bit_02_AUS3_STOP
   "Carrier_71_G120DControlWord.3" AT %I3910.3 : Bool;   // Bit_03_EN
   "Carrier_71_G120DControlWord.4" AT %I3910.4 : Bool;   // Bit_04_EN_RAMP
   "Carrier_71_G120DControlWord.5" AT %I3910.5 : Bool;   // Bit_05_START_RAMP
   "Carrier_71_G120DControlWord.6" AT %I3910.6 : Bool;   // Bit_06_SETPOINT
   "Carrier_71_G120DControlWord.7" AT %I3910.7 : Bool;   // Bit_07_RESET
   "Carrier_71_G120DControlWord.8" AT %I3911.0 : Bool;   // Bit_08_JOG_R
   "Carrier_71_G120DControlWord.9" AT %I3911.1 : Bool;   // Bit_09_JOG_L
   "Carrier_71_G120DControlWord.10" AT %I3911.2 : Bool;   // Bit_10_CONTR_PLC
   "Carrier_71_G120DControlWord.11" AT %I3911.3 : Bool;   // Bit_11_REVERSE
   "Carrier_71_G120DControlWord.12" AT %I3911.4 : Bool;   // Bit_12_BRAKE_RELEASE
   "Carrier_71_G120DControlWord.13" AT %I3911.5 : Bool;   // Bit_13_DDS
   "Carrier_71_G120DControlWord.14" AT %I3911.6 : Bool;   // Bit_14_DO0
   "Carrier_71_G120DControlWord.15" AT %I3911.7 : Bool;   // Bit_15_DO1
   "Carrier_71_G120DStatusWord" AT %IW3912 : Word;   // G120D_ZSW1_STATUS
   "Carrier_71_G120DStatusWord.0" AT %I3912.0 : Bool;   // Bit_00_READY_RUN
   "Carrier_71_G120DStatusWord.1" AT %I3912.1 : Bool;   // Bit_01_READY_ON
   "Carrier_71_G120DStatusWord.2" AT %I3912.2 : Bool;   // Bit_02_ENABLE
   "Carrier_71_G120DStatusWord.3" AT %I3912.3 : Bool;   // Bit_03_FAULT
   "Carrier_71_G120DStatusWord.4" AT %I3912.4 : Bool;   // Bit_04_OFF2
   "Carrier_71_G120DStatusWord.5" AT %I3912.5 : Bool;   // Bit_05_OFF3
   "Carrier_71_G120DStatusWord.6" AT %I3912.6 : Bool;   // Bit_06_LOCK_OUT
   "Carrier_71_G120DStatusWord.7" AT %I3912.7 : Bool;   // Bit_07_WARN
   "Carrier_71_G120DStatusWord.8" AT %I3913.0 : Bool;   // Bit_08_NO_DEVIATION
   "Carrier_71_G120DStatusWord.9" AT %I3913.1 : Bool;   // Bit_09_CONTR_PLC
   "Carrier_71_G120DStatusWord.10" AT %I3913.2 : Bool;   // Bit_10_F_MAX
   "Carrier_71_G120DStatusWord.11" AT %I3913.3 : Bool;   // Bit_11_LIMIT_REACHED
   "Carrier_71_G120DStatusWord.12" AT %I3913.4 : Bool;   // Bit_12_BRAKE_OPEN
   "Carrier_71_G120DStatusWord.13" AT %I3913.5 : Bool;   // Bit_13_NO_OVERTEMP
   "Carrier_71_G120DStatusWord.14" AT %I3913.6 : Bool;   // Bit_14_CW_CCW
   "Carrier_71_G120DStatusWord.15" AT %I3913.7 : Bool;   // Bit_15_OVERL
   "Carrier_71_Slot2_Input" AT %IW3914 : Word;   // SLOT 2 INPUT WORD
   "Carrier_71_CrashDetectSW" AT %I3914.0 : Bool;   // CRASH DETECT SW
   "Carrier_71_SpareSafetyInput(2_1)" AT %I3914.1 : Bool;   // SPARE SAFETY INPUT
   "Carrier_71_SpareSafetyInput(2_2)" AT %I3914.2 : Bool;   // SPARE SAFETY INPUT
   "Carrier_71_SpareSafetyInput(2_3)" AT %I3914.3 : Bool;   // SPARE SAFETY INPUT
   "Carrier_71_SpareSafetyInput(2_4)" AT %I3914.4 : Bool;   // SPARE SAFETY INPUT
   "Carrier_71_SpareSafetyInput(2_5)" AT %I3914.5 : Bool;   // SPARE SAFETY INPUT
   "Carrier_71_SpareSafetyInput(2_6)" AT %I3914.6 : Bool;   // SPARE SAFETY INPUT
   "Carrier_71_SpareSafetyInput(2_7)" AT %I3914.7 : Bool;   // SPARE SAFETY INPUT
   "Carrier_71_Slot3_SafetyOutput" AT %IW3915 : Word;   // SLOT 3 SAFETY OUTPUT WORD
   "Carrier_71_Crash_Detect_OK" AT %I3915.0 : Bool;   // CARRIER CRASH DETECT
   "Carrier_71_SpareSafetyOutput(3_1)" AT %I3915.1 : Bool;   // SPARE SAFETY OUTPUT
   "Carrier_71_SpareSafetyOutput(3_2)" AT %I3915.2 : Bool;   // SPARE SAFETY OUTPUT
   "Carrier_71_SpareSafetyOutput(3_3)" AT %I3915.3 : Bool;   // SPARE SAFETY OUTPUT
   "Carrier_71_SpareSafetyOutput(3_4)" AT %I3915.4 : Bool;   // SPARE SAFETY OUTPUT
   "Carrier_71_SpareSafetyOutput(3_5)" AT %I3915.5 : Bool;   // SPARE SAFETY OUTPUT
   "Carrier_71_SpareSafetyOutput(3_6)" AT %I3915.6 : Bool;   // SPARE SAFETY OUTPUT
   "Carrier_71_SpareSafetyOutput(3_7)" AT %I3915.7 : Bool;   // SPARE SAFETY OUTPUT
   "Carrier_71_Slot4_Input" AT %IW3916 : Word;   // SLOT 4 INPUT WORD
   "Carrier_71_480VPowerOn_MDCB1" AT %I3916.0 : Bool;   // 480 VAC POWER ON MDCB 1
   "Carrier_71_SpareInput(4_1)" AT %I3916.1 : Bool;   // SPARE INPUT
   "Carrier_71_SpareInput(4_2)" AT %I3916.2 : Bool;   // SPARE INPUT
   "Carrier_71_SitopSelectStatus" AT %I3916.3 : Bool;   // SITOP SELECT STATUS
   "Carrier_71_DCsupplyOnPSCB2" AT %I3916.4 : Bool;   // DC SUPPLY ON PSCB 2
   "Carrier_71_SpareInput(4_5)" AT %I3916.5 : Bool;   // SPARE INPUT
   "Carrier_71_SpareInput(4_6)" AT %I3916.6 : Bool;   // SPARE INPUT
   "Carrier_71_SpareInput(4_7)" AT %I3916.7 : Bool;   // SPARE INPUT
   "Carrier_71_PB1_ProdHoldLH" AT %I3917.0 : Bool;   // PB 1 PRODUCTION HOLD LH
   "Carrier_71_PB2_ResetLH" AT %I3917.1 : Bool;   // PB 2 RESET LH
   "Carrier_71_PB3_ProdHoldRH" AT %I3917.2 : Bool;   // PB 3 PRODUCTION HOLD RH
   "Carrier_71_PB4_ResetRH" AT %I3917.3 : Bool;   // PB 4 RESET RH
   "Carrier_71_SpareInput(4_14)" AT %I3917.4 : Bool;   // SPARE INPUT
   "Carrier_71_SpareInput(4_15)" AT %I3917.5 : Bool;   // SPARE INPUT
   "Carrier_71_SpareInput(4_16)" AT %I3917.6 : Bool;   // SPARE INPUT
   "Carrier_71_SpareInput(4_17)" AT %I3917.7 : Bool;   // SPARE INPUT
   "Carrier_71_Slot5_Output" AT %IW3918 : Word;   // SLOT 5 OUTPUT WORD
   "Carrier_71_IRD400_HMI_24VDC_ENABLE" AT %I3918.0 : Bool;   // IRD 400 PANEL HMI 24V DC POWER
   "Carrier_71_FaultLight_LH" AT %I3918.1 : Bool;   // FAULT LIGHT LH
   "Carrier_71_RunLight_LH" AT %I3918.2 : Bool;   // RUN LIGHT LH
   "Carrier_71_FaultLight_RH" AT %I3918.3 : Bool;   // FAULT LIGHT RH
   "Carrier_71_RunLight_RH" AT %I3918.4 : Bool;   // RUN LIGHT RH
   "Carrier_71_SpareOutput(5_5)" AT %I3918.5 : Bool;   // SPARE OUTPUT
   "Carrier_71_SpareOutput(5_6)" AT %I3918.6 : Bool;   // SPARE OUTPUT
   "Carrier_71_SpareOutput(5_7)" AT %I3918.7 : Bool;   // SPARE OUTPUT
   "Carrier_71_ActualSpeed" AT %IW3920 : Word;   // ACTUAL SPEED
   "Carrier_71_CarrierDriveAlarm" AT %IW3922 : Word;   // CARRIER DRIVE ALARM
   "Carrier_71_CarrierDriveWarning" AT %IW3924 : Word;   // CARRIER DRIVE WARNING
   "Carrier_72_Status" AT %IW3950 : Word;   // CARRIER STATUS WORD
   "Carrier_72_Status.0" AT %I3950.0 : Bool;   // HEARTBEAT
   "Carrier_72_Status.1" AT %I3950.1 : Bool;   // MANUAL
   "Carrier_72_Status.2" AT %I3950.2 : Bool;   // IN_AUTO
   "Carrier_72_Status.3" AT %I3950.3 : Bool;   // POSITIONING_COMPLETE
   "Carrier_72_Status.4" AT %I3950.4 : Bool;   // PRODUCTION HOLD
   "Carrier_72_Status.5" AT %I3950.5 : Bool;   // CARRIER MOVING FORWARD
   "Carrier_72_Status.6" AT %I3950.6 : Bool;   // CARRIER MOVING REVERSE
   "Carrier_72_Status.7" AT %I3950.7 : Bool;   // CARRIER FAULT
   "Carrier_72_Status.8" AT %I3951.0 : Bool;   // CRASH DETECT TRIPPED
   "Carrier_72_Status.9" AT %I3951.1 : Bool;
   "Carrier_72_Status.10" AT %I3951.2 : Bool;
   "Carrier_72_Status.11" AT %I3951.3 : Bool;
   "Carrier_72_Status.12" AT %I3951.4 : Bool;
   "Carrier_72_Status.13" AT %I3951.5 : Bool;
   "Carrier_72_Status.14" AT %I3951.6 : Bool;
   "Carrier_72_Status.15" AT %I3951.7 : Bool;
   "Carrier_72_SDCFaultCode" AT %IW3952 : Word;   // SDC FAULT CODE
   "Carrier_72_CarrierPosition" AT %ID3954 : DWord;   // CARRIER POSITION
   "Carrier_72_CarrierNumber" AT %IW3958 : Word;   // CARRIER NUMBER
   "Carrier_72_G120DControlWord" AT %IW3960 : Word;   // G120D_STW1_CONTROL
   "Carrier_72_G120DControlWord.0" AT %I3960.0 : Bool;   // Bit_00_ON
   "Carrier_72_G120DControlWord.1" AT %I3960.1 : Bool;   // Bit_01_AUS2_INH
   "Carrier_72_G120DControlWord.2" AT %I3960.2 : Bool;   // Bit_02_AUS3_STOP
   "Carrier_72_G120DControlWord.3" AT %I3960.3 : Bool;   // Bit_03_EN
   "Carrier_72_G120DControlWord.4" AT %I3960.4 : Bool;   // Bit_04_EN_RAMP
   "Carrier_72_G120DControlWord.5" AT %I3960.5 : Bool;   // Bit_05_START_RAMP
   "Carrier_72_G120DControlWord.6" AT %I3960.6 : Bool;   // Bit_06_SETPOINT
   "Carrier_72_G120DControlWord.7" AT %I3960.7 : Bool;   // Bit_07_RESET
   "Carrier_72_G120DControlWord.8" AT %I3961.0 : Bool;   // Bit_08_JOG_R
   "Carrier_72_G120DControlWord.9" AT %I3961.1 : Bool;   // Bit_09_JOG_L
   "Carrier_72_G120DControlWord.10" AT %I3961.2 : Bool;   // Bit_10_CONTR_PLC
   "Carrier_72_G120DControlWord.11" AT %I3961.3 : Bool;   // Bit_11_REVERSE
   "Carrier_72_G120DControlWord.12" AT %I3961.4 : Bool;   // Bit_12_BRAKE_RELEASE
   "Carrier_72_G120DControlWord.13" AT %I3961.5 : Bool;   // Bit_13_DDS